                           iReset := "DB2_WORK_BITS".Stacker_Handler.Input.iReset,
                           iAutomatic := "DB2_WORK_BITS".Stacker_Handler.Input.iAutomatic AND "Safe_S",
                           iManual := "DB2_WORK_BITS".Stacker_Handler.Input.iManual,
                           iManualUp := "O".CilindruVerticalStacker.ButAv,
                           iManualDown := "O".CilindruVerticalStacker.ButRet,
                           iManualOpenForks := "O".FurcaStacker.ButRet,
                           iManualCloseForks := "O".FurcaStacker.ButAv,
                           iB1_up := "DB2_WORK_BITS".Stacker_Handler.Input.Vertical_sus,
                           iB2_mid := "DB2_WORK_BITS".Stacker_Handler.Input.Vertical_mijloc,
                           iB10 := "DB2_WORK_BITS".Stacker_Handler.Input.iB10,
                           iB3_dwn := "DB2_WORK_BITS".Stacker_Handler.Input.Vertical_jos,
                           iB5_extins := "DB2_WORK_BITS".Stacker_Handler.Input.Furca_extins,
                           iB13_retras := "DB2_WORK_BITS".Stacker_Handler.Input.Furca_retras,
                           iB7_palet := "DB2_WORK_BITS".Stacker_Handler.Input.Detectie_palet,
                           iB8_stiva := "DB2_WORK_BITS".Stacker_Handler.Input.Senzor_stiva,
                           xSettings := "DB2_WORK_BITS".Settings_Stacker,
                           xHS_PalletDispencer := "DB2_WORK_BITS".Handshakes_Stacker,
                           oY4 => "DB2_WORK_BITS".Stacker_Handler.Output.Cmd_sus,
                           oY12 => "DB2_WORK_BITS".Stacker_Handler.Output.Cmd_jos,
                           oY6 => "DB2_WORK_BITS".Stacker_Handler.Output.Cmd_extindere,
                           oY14 => "DB2_WORK_BITS".Stacker_Handler.Output.Cmd_retragere,
                           oAlarmUpDown => "DB2_WORK_BITS".Stacker_Handler.Output.oAlarmUpDown,
                           oAlarmForks => "DB2_WORK_BITS".Stacker_Handler.Output.oAlarmForks,
                           oAlarmPosition => "DB2_WORK_BITS".Stacker_Handler.Output.oAlarmPosition,
                           oAlarmFull => "DB2_WORK_BITS".Stacker_Handler.Output.oAlarmFull,
                           ENO => #_w1);
   #dumyb := #_w1 AND "DB2_WORK_BITS".Stacker_Handler.Input.iEnable AND "DB2_WORK_BITS".Stacker_Handler.Input.iReset AND "DB2_WORK_BITS".Stacker_Handler.Input.iAutomatic AND "DB2_WORK_BITS".Stacker_Handler.Input.iAutomatic;
   IF #_w1 THEN #dumyw := "DB_PalletDispenser_PD2_Stacking_DB".PD1.Stepper; END_IF;
END_REGION

REGION Network 12: iEnable
   RUNG wire#powerrail
      Contact( "DB_MDM_S".Cycle_Run )
      wire#w1
      { S7_Templates := "SrcType := USInt" } NE_Contact(in1 := "s".f[4]."step", in2 := 8)
      Coil( "DB2_WORK_BITS".Stacker_Handler.Input.iEnable )
   END_RUNG
   RUNG wire#powerrail
      Contact( "DB_MDM_S".Manual )
   END_RUNG wire#w1
   RUNG wire#powerrail
      Contact( "DB_MDM_S".Init )
      wire#w2
      { S7_Templates := "SrcType := USInt" } EQ_Contact(in1 := "DB_Init_S"."step", in2 := 3)
   END_RUNG wire#w1
   RUNG wire#w2
      I_Contact( "b0" )
   END_RUNG wire#w1
   RUNG wire#powerrail
      Contact( "s".f[4].alm_disapear )
      Contact( "s".DeliveryStack )
      R_Coil( "DB2_WORK_BITS".Stacker_Handler.Input.iEnable )
   END_RUNG
   // the same network as SCL:
   "DB2_WORK_BITS".Stacker_Handler.Input.iEnable := ("DB_MDM_S".Cycle_Run OR "DB_MDM_S".Manual OR ("DB_MDM_S".Init AND (("DB_Init_S"."step" = 3) OR NOT "b0"))) AND ("s".f[4]."step" <> 8);
   IF "s".f[4].alm_disapear AND "s".DeliveryStack THEN
       "DB2_WORK_BITS".Stacker_Handler.Input.iEnable := FALSE;
   END_IF;
END_REGION

REGION Network 13: iAuto
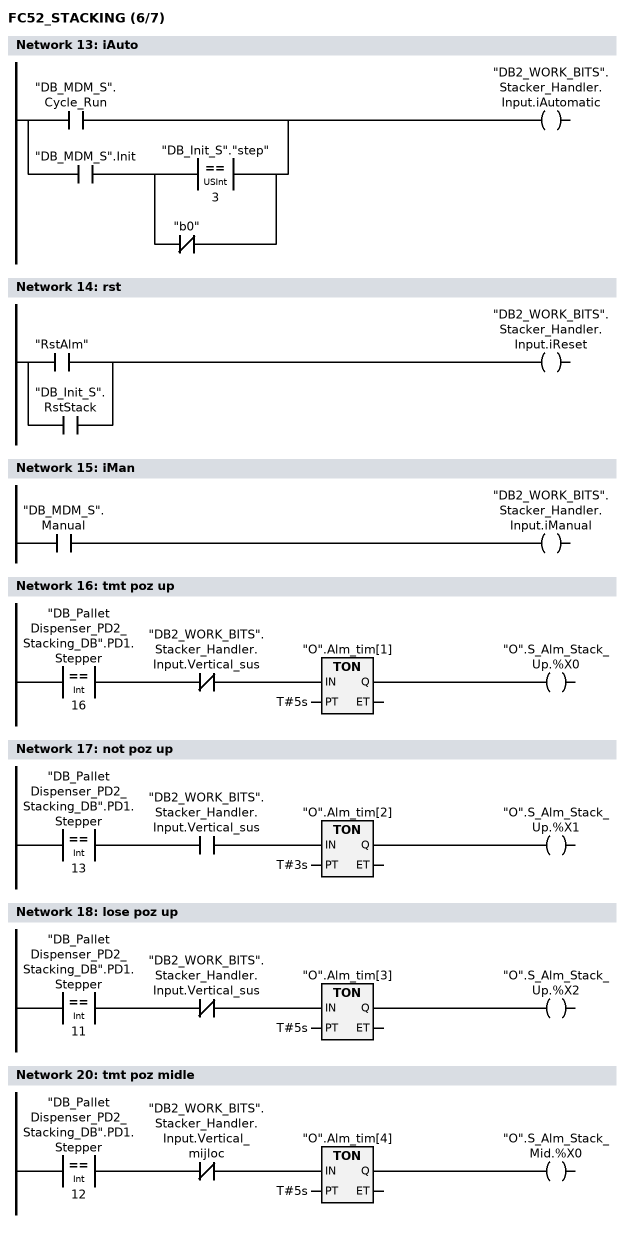
   RUNG wire#powerrail
      Contact( "DB_MDM_S".Cycle_Run )
      wire#w1
      Coil( "DB2_WORK_BITS".Stacker_Handler.Input.iAutomatic )
   END_RUNG
   RUNG wire#powerrail
      Contact( "DB_MDM_S".Init )
      wire#w2
      { S7_Templates := "SrcType := USInt" } EQ_Contact(in1 := "DB_Init_S"."step", in2 := 3)
   END_RUNG wire#w1
   RUNG wire#w2
      I_Contact( "b0" )
   END_RUNG wire#w1
   // the same network as SCL:
   "DB2_WORK_BITS".Stacker_Handler.Input.iAutomatic := "DB_MDM_S".Cycle_Run OR ("DB_MDM_S".Init AND (("DB_Init_S"."step" = 3) OR NOT "b0"));
END_REGION

REGION Network 14: rst
   RUNG wire#powerrail
      Contact( "RstAlm" )
      wire#w1
      Coil( "DB2_WORK_BITS".Stacker_Handler.Input.iReset )
   END_RUNG
   RUNG wire#powerrail
      Contact( "DB_Init_S".RstStack )
   END_RUNG wire#w1
   // the same network as SCL:
   "DB2_WORK_BITS".Stacker_Handler.Input.iReset := "RstAlm" OR "DB_Init_S".RstStack;
END_REGION

REGION Network 15: iMan
   RUNG wire#powerrail
      Contact( "DB_MDM_S".Manual )
      Coil( "DB2_WORK_BITS".Stacker_Handler.Input.iManual )
   END_RUNG
   // the same network as SCL:
   "DB2_WORK_BITS".Stacker_Handler.Input.iManual := "DB_MDM_S".Manual;
END_REGION

REGION Network 16: tmt poz up
   "O".Alm_tim[1].TON(IN := ("DB_PalletDispenser_PD2_Stacking_DB".PD1.Stepper = 16) AND NOT "DB2_WORK_BITS".Stacker_Handler.Input.Vertical_sus,
                      PT := T#5s);
   "O".S_Alm_Stack_Up.%X0 := "O".Alm_tim[1].Q;
END_REGION

REGION Network 17: not poz up
   "O".Alm_tim[2].TON(IN := ("DB_PalletDispenser_PD2_Stacking_DB".PD1.Stepper = 13) AND "DB2_WORK_BITS".Stacker_Handler.Input.Vertical_sus,
                      PT := T#3s);
   "O".S_Alm_Stack_Up.%X1 := "O".Alm_tim[2].Q;
END_REGION

REGION Network 18: lose poz up
   "O".Alm_tim[3].TON(IN := ("DB_PalletDispenser_PD2_Stacking_DB".PD1.Stepper = 11) AND NOT "DB2_WORK_BITS".Stacker_Handler.Input.Vertical_sus,
                      PT := T#5s);
   "O".S_Alm_Stack_Up.%X2 := "O".Alm_tim[3].Q;
END_REGION

REGION Network 19: lose poz up
END_REGION

REGION Network 20: tmt poz midle
   "O".Alm_tim[4].TON(IN := ("DB_PalletDispenser_PD2_Stacking_DB".PD1.Stepper = 12) AND NOT "DB2_WORK_BITS".Stacker_Handler.Input.Vertical_mijloc,
                      PT := T#5s);
   "O".S_Alm_Stack_Mid.%X0 := "O".Alm_tim[4].Q;
END_REGION

REGION Network 21: NoRls poz midle
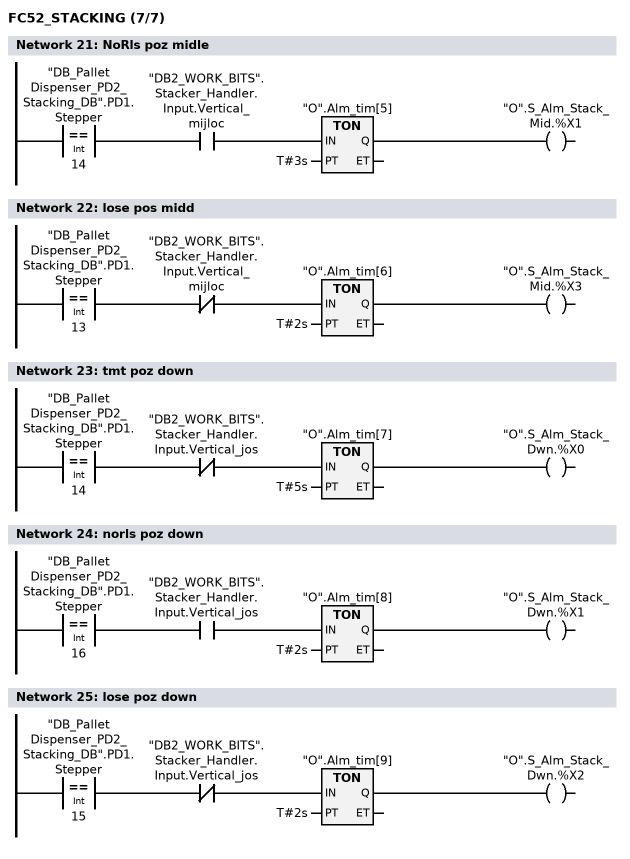
   "O".Alm_tim[5].TON(IN := ("DB_PalletDispenser_PD2_Stacking_DB".PD1.Stepper = 14) AND "DB2_WORK_BITS".Stacker_Handler.Input.Vertical_mijloc,
                      PT := T#3s);
   "O".S_Alm_Stack_Mid.%X1 := "O".Alm_tim[5].Q;
END_REGION

REGION Network 22: lose pos midd
   "O".Alm_tim[6].TON(IN := ("DB_PalletDispenser_PD2_Stacking_DB".PD1.Stepper = 13) AND NOT "DB2_WORK_BITS".Stacker_Handler.Input.Vertical_mijloc,
                      PT := T#2s);
   "O".S_Alm_Stack_Mid.%X3 := "O".Alm_tim[6].Q;
END_REGION

REGION Network 23: tmt poz down
   "O".Alm_tim[7].TON(IN := ("DB_PalletDispenser_PD2_Stacking_DB".PD1.Stepper = 14) AND NOT "DB2_WORK_BITS".Stacker_Handler.Input.Vertical_jos,
                      PT := T#5s);
   "O".S_Alm_Stack_Dwn.%X0 := "O".Alm_tim[7].Q;
END_REGION

REGION Network 24: norls poz down
   "O".Alm_tim[8].TON(IN := ("DB_PalletDispenser_PD2_Stacking_DB".PD1.Stepper = 16) AND "DB2_WORK_BITS".Stacker_Handler.Input.Vertical_jos,
                      PT := T#2s);
   "O".S_Alm_Stack_Dwn.%X1 := "O".Alm_tim[8].Q;
END_REGION

REGION Network 25: lose poz down
   "O".Alm_tim[9].TON(IN := ("DB_PalletDispenser_PD2_Stacking_DB".PD1.Stepper = 15) AND NOT "DB2_WORK_BITS".Stacker_Handler.Input.Vertical_jos,
                      PT := T#2s);
   "O".S_Alm_Stack_Dwn.%X2 := "O".Alm_tim[9].Q;
END_REGION
END_FUNCTION

FUNCTION "FC53_TRANSPORT_S" : Void   // FC53, LAD
{ S7_Optimized_Access := 'TRUE' }
VERSION : 0.1
   VAR_TEMP
      Transfer_Bit : Bool;
      SR_Down : Bool;
      SR_Out : Bool;
      DTR : Bool;
      Pallet_Centered : Bool;
      Send_to_Stacker : Bool;
      SQ_off : Bool;
      Send_bit : Bool;
      Finish_bit : Bool;
      Finish_Stack : Bool;
      Stacker_Basic : Bool;
      Send_Stack : Bool;
      Reset_counter : Bool;
      Reset_clock : Bool;
      P0_ON : Bool;
      P1_ON : Bool;
      P2_ON : Bool;
   END_VAR
   VAR_TEMP   // added for the SCL form of the ladder/FBD networks
      _w1 : Bool;
      _w2 : Bool;
      _w3 : Bool;
   END_VAR
BEGIN

REGION Network 1: centr
END_REGION

REGION Network 3
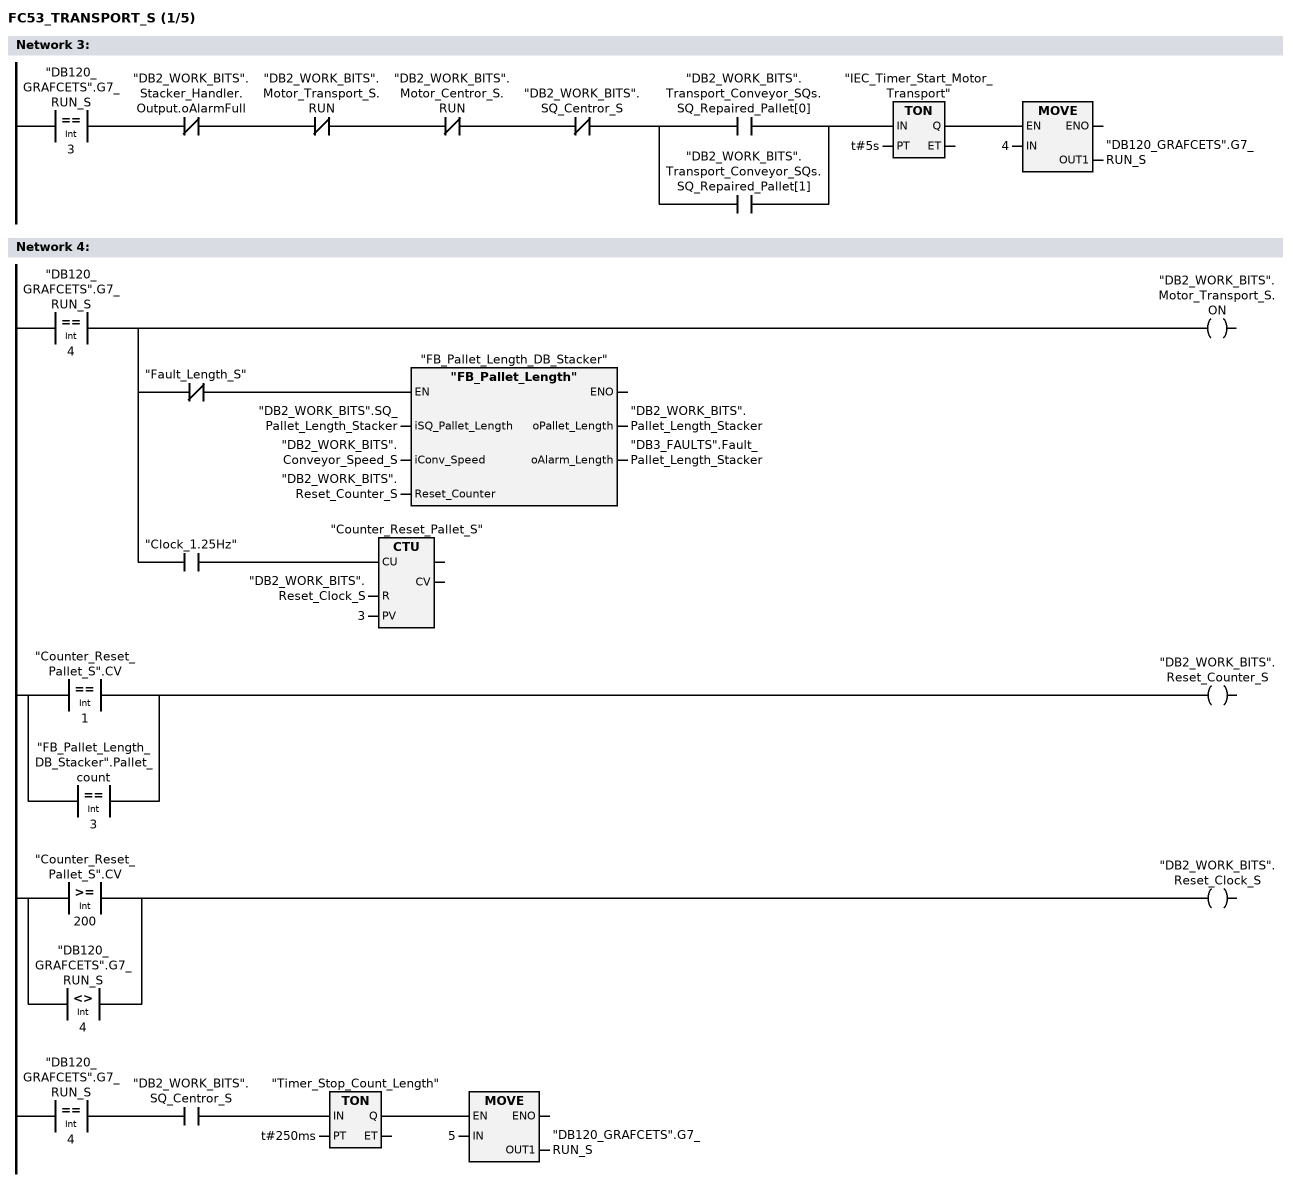
   "IEC_Timer_Start_Motor_Transport".TON(IN := ("DB120_GRAFCETS".G7_RUN_S = 3) AND NOT "DB2_WORK_BITS".Stacker_Handler.Output.oAlarmFull AND NOT "DB2_WORK_BITS".Motor_Transport_S.RUN AND NOT "DB2_WORK_BITS".Motor_Centror_S.RUN AND NOT "DB2_WORK_BITS".SQ_Centror_S AND ("DB2_WORK_BITS".Transport_Conveyor_SQs.SQ_Repaired_Pallet[0] OR "DB2_WORK_BITS".Transport_Conveyor_SQs.SQ_Repaired_Pallet[1]),
                           PT := t#5s);
   IF "IEC_Timer_Start_Motor_Transport".Q THEN "DB120_GRAFCETS".G7_RUN_S := 4; END_IF;
END_REGION

REGION Network 4
   "DB2_WORK_BITS".Motor_Transport_S.ON := "DB120_GRAFCETS".G7_RUN_S = 4;
   #_w1 := "DB2_WORK_BITS".Motor_Transport_S.ON;
   IF "DB2_WORK_BITS".Motor_Transport_S.ON AND NOT "Fault_Length_S" THEN
       "FB_Pallet_Length_DB_Stacker"(iSQ_Pallet_Length := "DB2_WORK_BITS".SQ_Pallet_Length_Stacker,   // "FB_Pallet_Length"
                               iConv_Speed := "DB2_WORK_BITS".Conveyor_Speed_S,
                               Reset_Counter := "DB2_WORK_BITS".Reset_Counter_S,
                               oPallet_Length => "DB2_WORK_BITS".Pallet_Length_Stacker,
                               oAlarm_Length => "DB3_FAULTS".Fault_Pallet_Length_Stacker);
   END_IF;
   "Counter_Reset_Pallet_S".CTU(CU := #_w1 AND "Clock_1.25Hz", R := "DB2_WORK_BITS".Reset_Clock_S, PV := 3);
   "DB2_WORK_BITS".Reset_Counter_S := ("Counter_Reset_Pallet_S".CV = 1) OR ("FB_Pallet_Length_DB_Stacker".Pallet_count = 3);
   "DB2_WORK_BITS".Reset_Clock_S := ("Counter_Reset_Pallet_S".CV >= 200) OR ("DB120_GRAFCETS".G7_RUN_S <> 4);
   "Timer_Stop_Count_Length".TON(IN := ("DB120_GRAFCETS".G7_RUN_S = 4) AND "DB2_WORK_BITS".SQ_Centror_S,
                           PT := t#250ms);
   IF "Timer_Stop_Count_Length".Q THEN "DB120_GRAFCETS".G7_RUN_S := 5; END_IF;
END_REGION

REGION Network 5
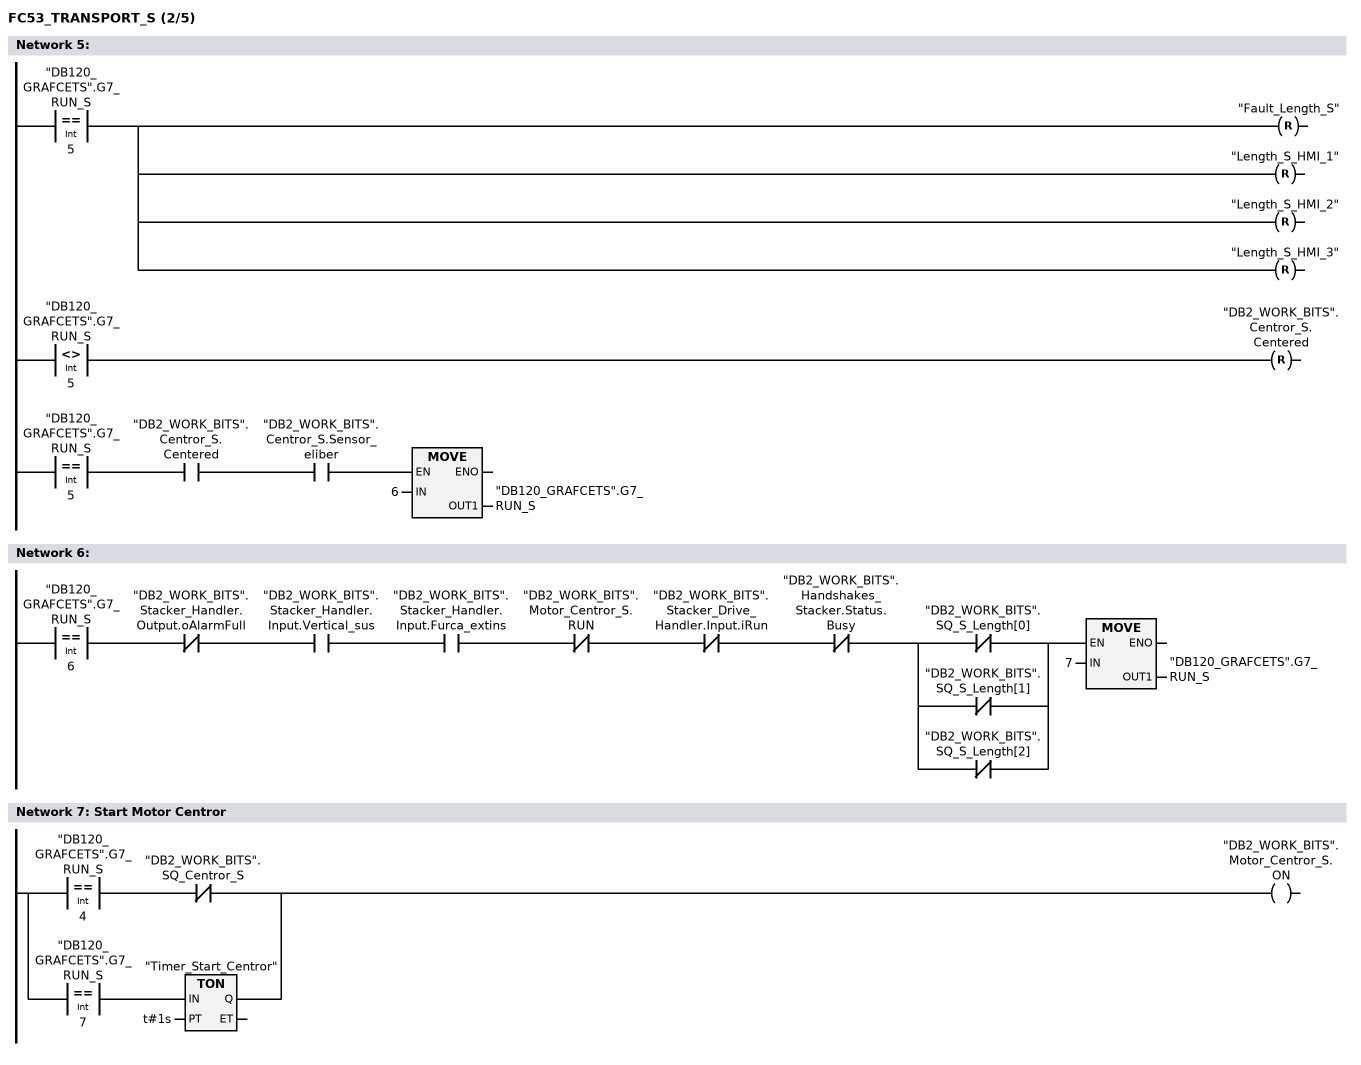
   RUNG wire#powerrail
      { S7_Templates := "SrcType := Int" } EQ_Contact(in1 := "DB120_GRAFCETS".G7_RUN_S, in2 := 5)
      wire#w1
      R_Coil( "Fault_Length_S" )
   END_RUNG
   RUNG wire#w1
      R_Coil( "Length_S_HMI_1" )
   END_RUNG
   RUNG wire#w1
      R_Coil( "Length_S_HMI_2" )
   END_RUNG
   RUNG wire#w1
      R_Coil( "Length_S_HMI_3" )
   END_RUNG
   RUNG wire#powerrail
      { S7_Templates := "SrcType := Int" } NE_Contact(in1 := "DB120_GRAFCETS".G7_RUN_S, in2 := 5)
      R_Coil( "DB2_WORK_BITS".Centror_S.Centered )
   END_RUNG
   RUNG wire#powerrail
      { S7_Templates := "SrcType := Int" } EQ_Contact(in1 := "DB120_GRAFCETS".G7_RUN_S, in2 := 5)
      Contact( "DB2_WORK_BITS".Centror_S.Centered )
      Contact( "DB2_WORK_BITS".Centror_S.Sensor_eliber )
      Move(in := 6, out1 => "DB120_GRAFCETS".G7_RUN_S)
   END_RUNG
   // the same network as SCL:
   IF "DB120_GRAFCETS".G7_RUN_S = 5 THEN
       "Fault_Length_S" := FALSE;
       "Length_S_HMI_1" := FALSE;
       "Length_S_HMI_2" := FALSE;
       "Length_S_HMI_3" := FALSE;
   END_IF;
   IF "DB120_GRAFCETS".G7_RUN_S <> 5 THEN "DB2_WORK_BITS".Centror_S.Centered := FALSE; END_IF;
   IF ("DB120_GRAFCETS".G7_RUN_S = 5) AND "DB2_WORK_BITS".Centror_S.Centered AND "DB2_WORK_BITS".Centror_S.Sensor_eliber THEN
       "DB120_GRAFCETS".G7_RUN_S := 6;
   END_IF;
END_REGION

REGION Network 6
   RUNG wire#powerrail
      { S7_Templates := "SrcType := Int" } EQ_Contact(in1 := "DB120_GRAFCETS".G7_RUN_S, in2 := 6)
      I_Contact( "DB2_WORK_BITS".Stacker_Handler.Output.oAlarmFull )
      Contact( "DB2_WORK_BITS".Stacker_Handler.Input.Vertical_sus )
      Contact( "DB2_WORK_BITS".Stacker_Handler.Input.Furca_extins )
      I_Contact( "DB2_WORK_BITS".Motor_Centror_S.RUN )
      I_Contact( "DB2_WORK_BITS".Stacker_Drive_Handler.Input.iRun )
      I_Contact( "DB2_WORK_BITS".Handshakes_Stacker.Status.Busy )
      wire#w1
      I_Contact( "DB2_WORK_BITS".SQ_S_Length[0] )
      wire#w2
      Move(in := 7, out1 => "DB120_GRAFCETS".G7_RUN_S)
   END_RUNG
   RUNG wire#w1
      I_Contact( "DB2_WORK_BITS".SQ_S_Length[1] )
   END_RUNG wire#w2
   RUNG wire#w1
      I_Contact( "DB2_WORK_BITS".SQ_S_Length[2] )
   END_RUNG wire#w2
   // the same network as SCL:
   IF ("DB120_GRAFCETS".G7_RUN_S = 6) AND NOT "DB2_WORK_BITS".Stacker_Handler.Output.oAlarmFull AND "DB2_WORK_BITS".Stacker_Handler.Input.Vertical_sus AND "DB2_WORK_BITS".Stacker_Handler.Input.Furca_extins AND NOT "DB2_WORK_BITS".Motor_Centror_S.RUN AND NOT "DB2_WORK_BITS".Stacker_Drive_Handler.Input.iRun AND NOT "DB2_WORK_BITS".Handshakes_Stacker.Status.Busy AND (NOT "DB2_WORK_BITS".SQ_S_Length[0] OR NOT "DB2_WORK_BITS".SQ_S_Length[1] OR NOT "DB2_WORK_BITS".SQ_S_Length[2]) THEN
       "DB120_GRAFCETS".G7_RUN_S := 7;
   END_IF;
END_REGION

REGION Network 7: Start Motor Centror
   "Timer_Start_Centror".TON(IN := "DB120_GRAFCETS".G7_RUN_S = 7, PT := t#1s);
   "DB2_WORK_BITS".Motor_Centror_S.ON := (("DB120_GRAFCETS".G7_RUN_S = 4) AND NOT "DB2_WORK_BITS".SQ_Centror_S) OR "Timer_Start_Centror".Q;
END_REGION

REGION Network 8: Start Motor Stacker
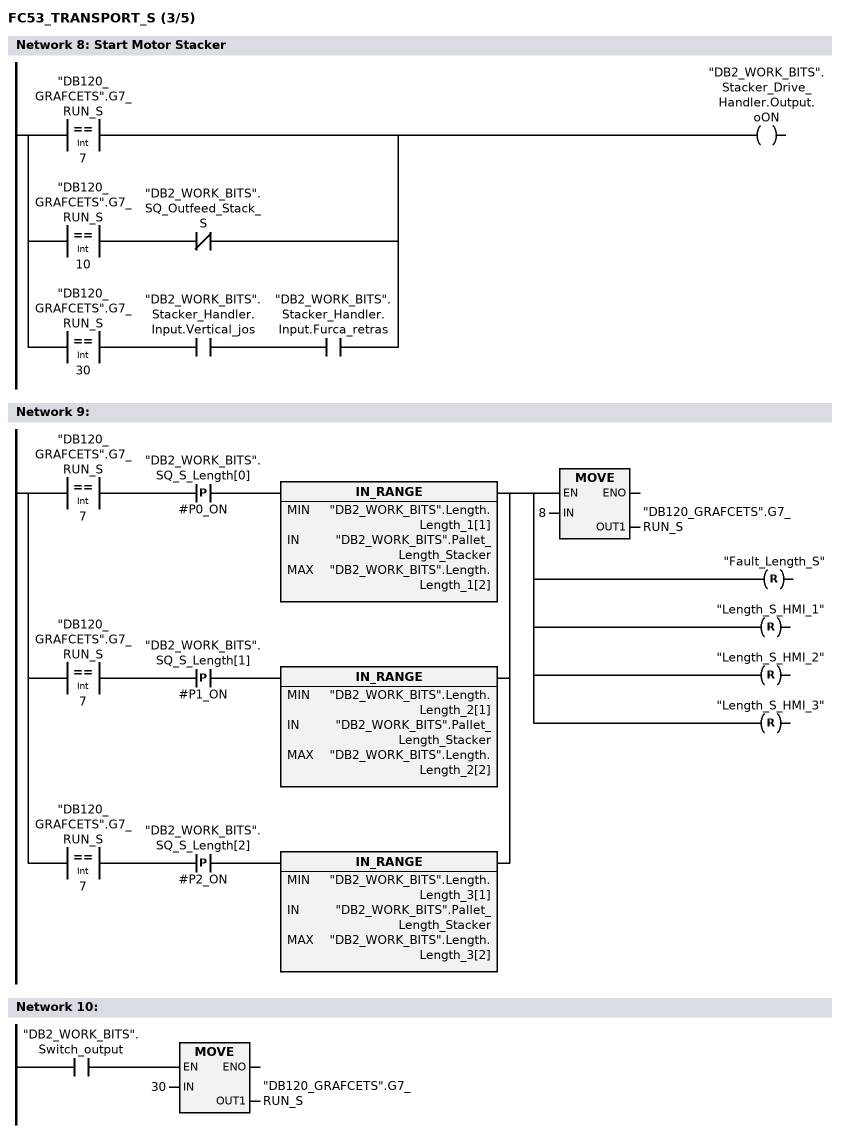
   RUNG wire#powerrail
      { S7_Templates := "SrcType := Int" } EQ_Contact(in1 := "DB120_GRAFCETS".G7_RUN_S, in2 := 7)
      wire#w1
      Coil( "DB2_WORK_BITS".Stacker_Drive_Handler.Output.oON )
   END_RUNG
   RUNG wire#powerrail
      { S7_Templates := "SrcType := Int" } EQ_Contact(in1 := "DB120_GRAFCETS".G7_RUN_S, in2 := 10)
      I_Contact( "DB2_WORK_BITS".SQ_Outfeed_Stack_S )
   END_RUNG wire#w1
   RUNG wire#powerrail
      { S7_Templates := "SrcType := Int" } EQ_Contact(in1 := "DB120_GRAFCETS".G7_RUN_S, in2 := 30)
      Contact( "DB2_WORK_BITS".Stacker_Handler.Input.Vertical_jos )
      Contact( "DB2_WORK_BITS".Stacker_Handler.Input.Furca_retras )
   END_RUNG wire#w1
   // the same network as SCL:
   "DB2_WORK_BITS".Stacker_Drive_Handler.Output.oON := ("DB120_GRAFCETS".G7_RUN_S = 7) OR (("DB120_GRAFCETS".G7_RUN_S = 10) AND NOT "DB2_WORK_BITS".SQ_Outfeed_Stack_S) OR (("DB120_GRAFCETS".G7_RUN_S = 30) AND "DB2_WORK_BITS".Stacker_Handler.Input.Vertical_jos AND "DB2_WORK_BITS".Stacker_Handler.Input.Furca_retras);
END_REGION

REGION Network 9
   RUNG wire#powerrail
      { S7_Templates := "SrcType := Int" } EQ_Contact(in1 := "DB120_GRAFCETS".G7_RUN_S, in2 := 7)
      P_Contact(operand := "DB2_WORK_BITS".SQ_S_Length[0], bit := #P0_ON)
      { S7_Templates := "SrcType := Int" } InRange(min := "DB2_WORK_BITS".Length.Length_1[1], in := "DB2_WORK_BITS".Pallet_Length_Stacker, max := "DB2_WORK_BITS".Length.Length_1[2])
      wire#w1
      Move(in := 8, out1 => "DB120_GRAFCETS".G7_RUN_S)
   END_RUNG
   RUNG wire#powerrail
      { S7_Templates := "SrcType := Int" } EQ_Contact(in1 := "DB120_GRAFCETS".G7_RUN_S, in2 := 7)
      P_Contact(operand := "DB2_WORK_BITS".SQ_S_Length[1], bit := #P1_ON)
      { S7_Templates := "SrcType := Int" } InRange(min := "DB2_WORK_BITS".Length.Length_2[1], in := "DB2_WORK_BITS".Pallet_Length_Stacker, max := "DB2_WORK_BITS".Length.Length_2[2])
   END_RUNG wire#w1
   RUNG wire#powerrail
      { S7_Templates := "SrcType := Int" } EQ_Contact(in1 := "DB120_GRAFCETS".G7_RUN_S, in2 := 7)
      P_Contact(operand := "DB2_WORK_BITS".SQ_S_Length[2], bit := #P2_ON)
      { S7_Templates := "SrcType := Int" } InRange(min := "DB2_WORK_BITS".Length.Length_3[1], in := "DB2_WORK_BITS".Pallet_Length_Stacker, max := "DB2_WORK_BITS".Length.Length_3[2])
   END_RUNG wire#w1
   RUNG wire#w1
      R_Coil( "Fault_Length_S" )
   END_RUNG
   RUNG wire#w1
      R_Coil( "Length_S_HMI_1" )
   END_RUNG
   RUNG wire#w1
      R_Coil( "Length_S_HMI_2" )
   END_RUNG
   RUNG wire#w1
      R_Coil( "Length_S_HMI_3" )
   END_RUNG
   // the same network as SCL:
   #_w1 := ("DB120_GRAFCETS".G7_RUN_S = 7) AND "DB2_WORK_BITS".SQ_S_Length[0] AND NOT #P0_ON;   // rising edge of "DB2_WORK_BITS".SQ_S_Length[0]
   #P0_ON := "DB2_WORK_BITS".SQ_S_Length[0];
   #_w2 := ("DB120_GRAFCETS".G7_RUN_S = 7) AND "DB2_WORK_BITS".SQ_S_Length[1] AND NOT #P1_ON;   // rising edge of "DB2_WORK_BITS".SQ_S_Length[1]
   #P1_ON := "DB2_WORK_BITS".SQ_S_Length[1];
   #_w3 := ("DB120_GRAFCETS".G7_RUN_S = 7) AND "DB2_WORK_BITS".SQ_S_Length[2] AND NOT #P2_ON;   // rising edge of "DB2_WORK_BITS".SQ_S_Length[2]
   #P2_ON := "DB2_WORK_BITS".SQ_S_Length[2];
   IF (#_w1 AND ("DB2_WORK_BITS".Length.Length_1[1] <= "DB2_WORK_BITS".Pallet_Length_Stacker) AND ("DB2_WORK_BITS".Pallet_Length_Stacker <= "DB2_WORK_BITS".Length.Length_1[2])) OR (#_w2 AND ("DB2_WORK_BITS".Length.Length_2[1] <= "DB2_WORK_BITS".Pallet_Length_Stacker) AND ("DB2_WORK_BITS".Pallet_Length_Stacker <= "DB2_WORK_BITS".Length.Length_2[2])) OR (#_w3 AND ("DB2_WORK_BITS".Length.Length_3[1] <= "DB2_WORK_BITS".Pallet_Length_Stacker) AND ("DB2_WORK_BITS".Pallet_Length_Stacker <= "DB2_WORK_BITS".Length.Length_3[2])) THEN
       "DB120_GRAFCETS".G7_RUN_S := 8;
       "Fault_Length_S" := FALSE;
       "Length_S_HMI_1" := FALSE;
       "Length_S_HMI_2" := FALSE;
       "Length_S_HMI_3" := FALSE;
   END_IF;
END_REGION

REGION Network 10
   RUNG wire#powerrail
      Contact( "DB2_WORK_BITS".Switch_output )
      Move(in := 30, out1 => "DB120_GRAFCETS".G7_RUN_S)
   END_RUNG
   // the same network as SCL:
   IF "DB2_WORK_BITS".Switch_output THEN "DB120_GRAFCETS".G7_RUN_S := 30; END_IF;
END_REGION

REGION Network 11
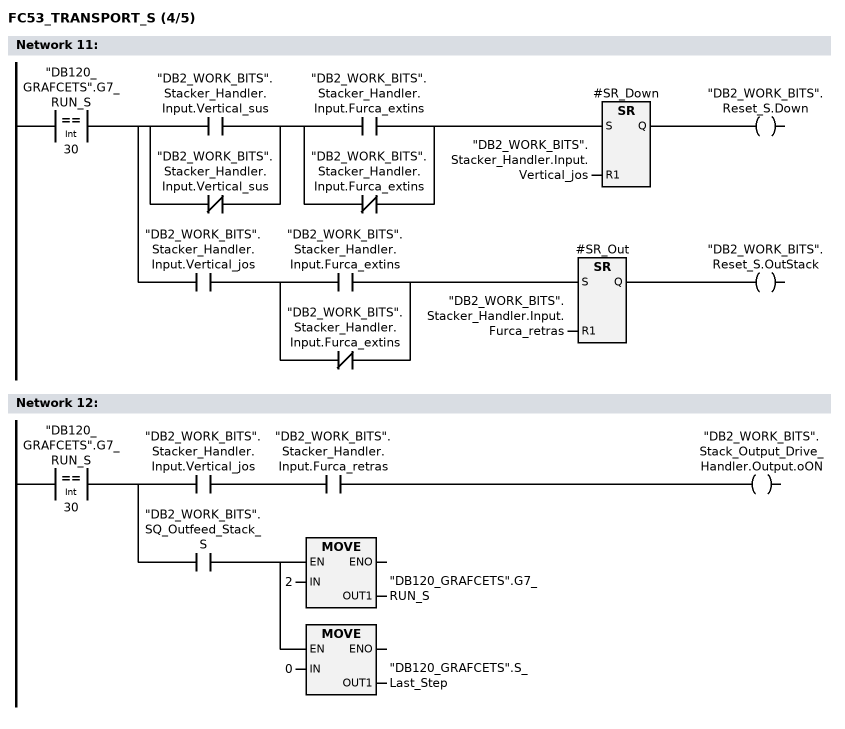
   RUNG wire#powerrail
      { S7_Templates := "SrcType := Int" } EQ_Contact(in1 := "DB120_GRAFCETS".G7_RUN_S, in2 := 30)
      wire#w1
      Contact( "DB2_WORK_BITS".Stacker_Handler.Input.Vertical_sus )
      wire#w2
      Contact( "DB2_WORK_BITS".Stacker_Handler.Input.Furca_extins )
      wire#w3
      S_SR(operand := #SR_Down, r1 := "DB2_WORK_BITS".Stacker_Handler.Input.Vertical_jos)
      Coil( "DB2_WORK_BITS".Reset_S.Down )
   END_RUNG
   RUNG wire#w1
      I_Contact( "DB2_WORK_BITS".Stacker_Handler.Input.Vertical_sus )
   END_RUNG wire#w2
   RUNG wire#w2
      I_Contact( "DB2_WORK_BITS".Stacker_Handler.Input.Furca_extins )
   END_RUNG wire#w3
   RUNG wire#w1
      Contact( "DB2_WORK_BITS".Stacker_Handler.Input.Vertical_jos )
      wire#w4
      Contact( "DB2_WORK_BITS".Stacker_Handler.Input.Furca_extins )
      wire#w5
      S_SR(operand := #SR_Out, r1 := "DB2_WORK_BITS".Stacker_Handler.Input.Furca_retras)
      Coil( "DB2_WORK_BITS".Reset_S.OutStack )
   END_RUNG
   RUNG wire#w4
      I_Contact( "DB2_WORK_BITS".Stacker_Handler.Input.Furca_extins )
   END_RUNG wire#w5
   // the same network as SCL:
   #_w1 := "DB120_GRAFCETS".G7_RUN_S = 30;
   IF #_w1 AND ("DB2_WORK_BITS".Stacker_Handler.Input.Vertical_sus OR NOT "DB2_WORK_BITS".Stacker_Handler.Input.Vertical_sus) AND ("DB2_WORK_BITS".Stacker_Handler.Input.Furca_extins OR NOT "DB2_WORK_BITS".Stacker_Handler.Input.Furca_extins) THEN
       #SR_Down := TRUE;   // SR flip-flop
   END_IF;
   IF "DB2_WORK_BITS".Stacker_Handler.Input.Vertical_jos THEN #SR_Down := FALSE; END_IF;
   "DB2_WORK_BITS".Reset_S.Down := #SR_Down;
   IF #_w1 AND "DB2_WORK_BITS".Stacker_Handler.Input.Vertical_jos AND ("DB2_WORK_BITS".Stacker_Handler.Input.Furca_extins OR NOT "DB2_WORK_BITS".Stacker_Handler.Input.Furca_extins) THEN
       #SR_Out := TRUE;   // SR flip-flop
   END_IF;
   IF "DB2_WORK_BITS".Stacker_Handler.Input.Furca_retras THEN #SR_Out := FALSE; END_IF;
   "DB2_WORK_BITS".Reset_S.OutStack := #SR_Out;
END_REGION

REGION Network 12
   RUNG wire#powerrail
      { S7_Templates := "SrcType := Int" } EQ_Contact(in1 := "DB120_GRAFCETS".G7_RUN_S, in2 := 30)
      wire#w1
      Contact( "DB2_WORK_BITS".Stacker_Handler.Input.Vertical_jos )
      Contact( "DB2_WORK_BITS".Stacker_Handler.Input.Furca_retras )
      Coil( "DB2_WORK_BITS".Stack_Output_Drive_Handler.Output.oON )
   END_RUNG
   RUNG wire#w1
      Contact( "DB2_WORK_BITS".SQ_Outfeed_Stack_S )
      wire#w2
      Move(in := 2, out1 => "DB120_GRAFCETS".G7_RUN_S)
   END_RUNG
   RUNG wire#w2
      Move(in := 0, out1 => "DB120_GRAFCETS".S_Last_Step)
   END_RUNG
   // the same network as SCL:
   #_w1 := "DB120_GRAFCETS".G7_RUN_S = 30;
   "DB2_WORK_BITS".Stack_Output_Drive_Handler.Output.oON := #_w1 AND "DB2_WORK_BITS".Stacker_Handler.Input.Vertical_jos AND "DB2_WORK_BITS".Stacker_Handler.Input.Furca_retras;
   IF #_w1 AND "DB2_WORK_BITS".SQ_Outfeed_Stack_S THEN
       "DB120_GRAFCETS".G7_RUN_S := 2;
       "DB120_GRAFCETS".S_Last_Step := 0;
   END_IF;
END_REGION

REGION Network 13: Fault Length S
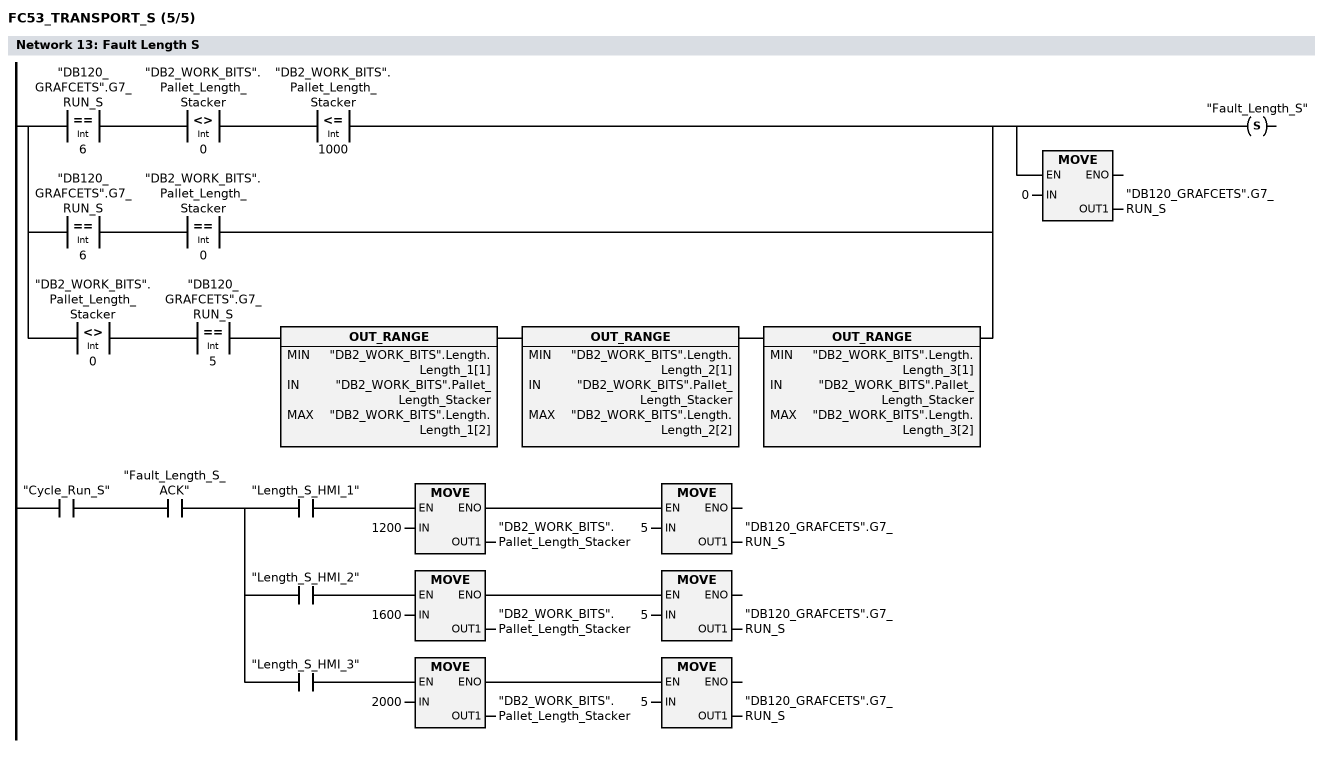
   IF (("DB120_GRAFCETS".G7_RUN_S = 6) AND ("DB2_WORK_BITS".Pallet_Length_Stacker <> 0) AND ("DB2_WORK_BITS".Pallet_Length_Stacker <= 1000)) OR (("DB120_GRAFCETS".G7_RUN_S = 6) AND ("DB2_WORK_BITS".Pallet_Length_Stacker = 0)) OR (("DB2_WORK_BITS".Pallet_Length_Stacker <> 0) AND ("DB120_GRAFCETS".G7_RUN_S = 5) AND (("DB2_WORK_BITS".Pallet_Length_Stacker < "DB2_WORK_BITS".Length.Length_1[1]) OR ("DB2_WORK_BITS".Pallet_Length_Stacker > "DB2_WORK_BITS".Length.Length_1[2])) AND (("DB2_WORK_BITS".Pallet_Length_Stacker < "DB2_WORK_BITS".Length.Length_2[1]) OR ("DB2_WORK_BITS".Pallet_Length_Stacker > "DB2_WORK_BITS".Length.Length_2[2])) AND (("DB2_WORK_BITS".Pallet_Length_Stacker < "DB2_WORK_BITS".Length.Length_3[1]) OR ("DB2_WORK_BITS".Pallet_Length_Stacker > "DB2_WORK_BITS".Length.Length_3[2]))) THEN
       "Fault_Length_S" := TRUE;
       "DB120_GRAFCETS".G7_RUN_S := 0;
   END_IF;
   #_w1 := "Cycle_Run_S" AND "Fault_Length_S_ACK";
   IF #_w1 AND "Length_S_HMI_1" THEN
       "DB2_WORK_BITS".Pallet_Length_Stacker := 1200;
       "DB120_GRAFCETS".G7_RUN_S := 5;
   END_IF;
   IF #_w1 AND "Length_S_HMI_2" THEN
       "DB2_WORK_BITS".Pallet_Length_Stacker := 1600;
       "DB120_GRAFCETS".G7_RUN_S := 5;
   END_IF;
   IF #_w1 AND "Length_S_HMI_3" THEN
       "DB2_WORK_BITS".Pallet_Length_Stacker := 2000;
       "DB120_GRAFCETS".G7_RUN_S := 5;
   END_IF;
END_REGION
END_FUNCTION

FUNCTION "FC55_MAINTENANCE_1" : Void   // FC55, LAD
{ S7_Optimized_Access := 'TRUE' }
VERSION : 0.1
BEGIN

REGION Network 1